(* Logix 5000 project; controller MV vendor 1 type 14 code 217 rev 31.11; software revision 31.00; part 11 of 53 *)
(* tags used below, declared in another part *)
   MC_CIP_String_Result1 : DINT;
   MC_CIP_String_Result2 : DINT;
   MC_CIP_String_Result3 : DINT;
   MC_CIP_String_Result4 : DINT;
   MC_CIP_String_Result5 : DINT;
   MC_CIP_String_Result6 : DINT;
   BH_Draindown_ON : DINT;
   CWD : CHECKWORD_FLAGS;
   FRHR26_31_Valves_ON_Produced : DINT;
   FVHR12_1701 : PlantItem;   // Valve FVHR12_17/01
   FVHR12_1702 : PlantItem;   // Valve FVHR12_17/02
   FVHR12_1703 : PlantItem;   // Valve FVHR12_17/03
   FVHR12_17_Valves_ON : BOOL;   // Check bit to confirm valves for FV12-17 route are open
   FVHR18_21_Valves_ON : BOOL;   // Check bit to confirm valves for FV18-21 route are open
   FVHR18_2501 : PlantItem;   // Valve FVHR18_25/01
   FVHR18_2502 : PlantItem;   // Valve FVHR18_25/02
   FVHR18_2503 : PlantItem;   // Valve FVHR18_25/03
   FVHR18_2504 : PlantItem;   // Valve FVHR18_25/04
   FVHR18_2505 : PlantItem;   // Valve FVHR18_25/05
   FVHR18_2506 : PlantItem;   // Valve FVHR18_25/06
   FVHR1_1101 : PlantItem;   // Valve FVHR1_11/01
   FVHR1_1102 : PlantItem;   // Valve FVHR1_11/02
   FVHR1_1103 : PlantItem;   // Valve FVHR1_11/03
   FVHR1_11_Valves_ON : BOOL;   // Check bit to confirm valves for FV1-11 route are open
   FVHR1_1701 : PlantItem;   // Valve FVHR1_17/01
   FVHR22_25_Valves_ON : BOOL;   // Check bit to confirm valves for FV22-25 route are open
   FVHR26_3101 : PlantItem;   // Valve FVHR26_31/01
   FVHR26_3102 : PlantItem;   // Valve FVHR26_31/02
   FVHR26_3103 : PlantItem;   // Valve FVHR26_31/03
   FVHR26_31_Valves_ON : BOOL;   // Check bit to confirm valves for FV26-31 route are open
   FVHRLTX02_IP : PlantItem;   // Effluent Tank Level Transmitter
   FVHRM02 : PlantItem;   // Valve FVHRM02
   FVHRM03 : PlantItem;   // Valve FVHRM03
   FVHRM04 : PlantItem;   // Valve FVHRM04
   FVHRMD01 : PlantItem;   // Valve FVHRMD01
   FVHRTM01_IP : PlantItem;   // Turbidty Meter FVHRTM01
   IGI_TestBit : BOOL;
   MC_bit_returned : BOOL;
   MC_CH2_CIP_BYPASS_Conditions : BOOL;
   MC_CH2_CIP_BYPASS_DrainConditions : BOOL;
   MC_CH2_CIP_Messages : STRING[20];   // CH2 CIP Scada Messages
   MC_CH2_CIP_YST_Scb_Bypass : BOOL;
   MC_CH2_DR1 : PlantItem;   // CH2_DR1
   MC_CH2_DR2 : PlantItem;   // CH2_DR2
   MC_CH2_DT1 : PlantItem;   // CH2_DT1
   MC_CH2_DT2 : PlantItem;   // CH2_DT2
   MC_CH2_FVBypass_Flush_ALARM : ALARM_DIGITAL;
   MC_CH2_FVBYPASS_H2O_Flush : BOOL;
   MC_CH2_R1 : PlantItem;   // CH2_R1
   MC_CH2_R1R : PlantItem;   // CH2_R1R
   MC_CH2_R2 : PlantItem;   // CH2_R2
   MC_CH2_R2R : PlantItem;   // CH2_R2R
   MC_CH2_R3 : PlantItem;   // CH2_R3
   MC_CH2_R3R : PlantItem;   // CH2_R3R
   MC_CH2_R4 : PlantItem;   // CH2_R4
   MC_CH2_R4R : PlantItem;   // CH2_R4R
   MC_CH2_R5 : PlantItem;   // CH2_R5
   MC_CH2_R5R : PlantItem;   // CH2_R5R
   MC_CH2_R6 : PlantItem;   // CH2_R6
   MC_CH2_R6R : PlantItem;   // CH2_R6R
   MC_CH2_TURBID_High : BOOL;
   MC_CIP_CH2_String_OK : BOOL;
   MC_CIP_CH2_Strings_HopRinse : STRING[30];
   MC_CIP_EFFTank_Full : BOOL;
   MC_CIP_EFFTank_Start_Lvl_Ok : BOOL;
   MC_N10 : INT[255];   // SETTINGS
   MC_N112 : INT[255];   // FVR DATA Data read from FV ro uting PLC
   MC_N113 : INT[255];   // MVR DATA Data read from MV ro uting PLC
   MC_N114 : INT[255];   // YP DATA
   MC_N120 : INT[255];   // C2 PLC Channel 2 PLC data
   MC_N122 : INT[255];   // CH2 PROG Channel 2 CIP progra m
   MC_N200 : INT[255];   // CHK_WORK Plant item fault che cking work area
   MC_N7 : INT[255];   // INTEGER
   MC_P2 : PlantItem;   // P2
   MC_PX_100 : PlantItem;   // PX_100
   MC_PX_101 : PlantItem;   // PX_101
   MC_T125 : TIMER[255];   // CH2 TIMERS Channel 2 timers
   MC_T4 : TIMER[255];   // TIMER
(* MC_Common, continued *)

ROUTINE MC_CH2_GLOBL_125   (* ladder *)
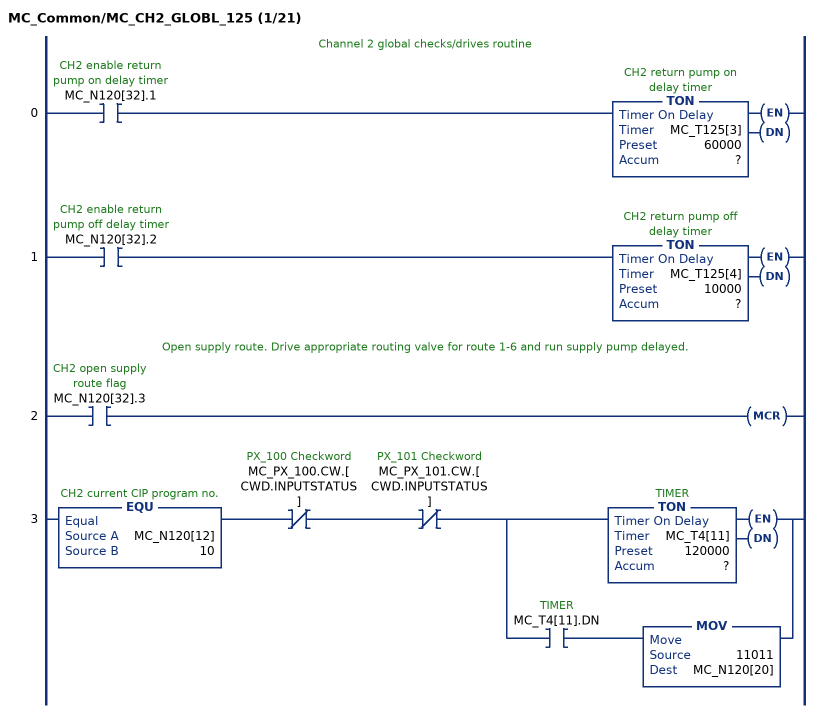
   // Channel 2 global checks/drives routine
   0: XIC(MC_N120[32].1)TON(MC_T125[3],?,?);
   1: XIC(MC_N120[32].2)TON(MC_T125[4],?,?);
   // Open supply route. Drive appropriate routing valve for route 1-6 and run supply pump delayed.
   2: XIC(MC_N120[32].3)MCR();
   3: EQU(MC_N120[12],10)XIO(MC_PX_100.CW.[CWD.INPUTSTATUS])XIO(MC_PX_101.CW.[CWD.INPUTSTATUS])[TON(MC_T4[11],?,?) ,XIC(MC_T4[11].DN) MOV(11011,MC_N120[20]) ];
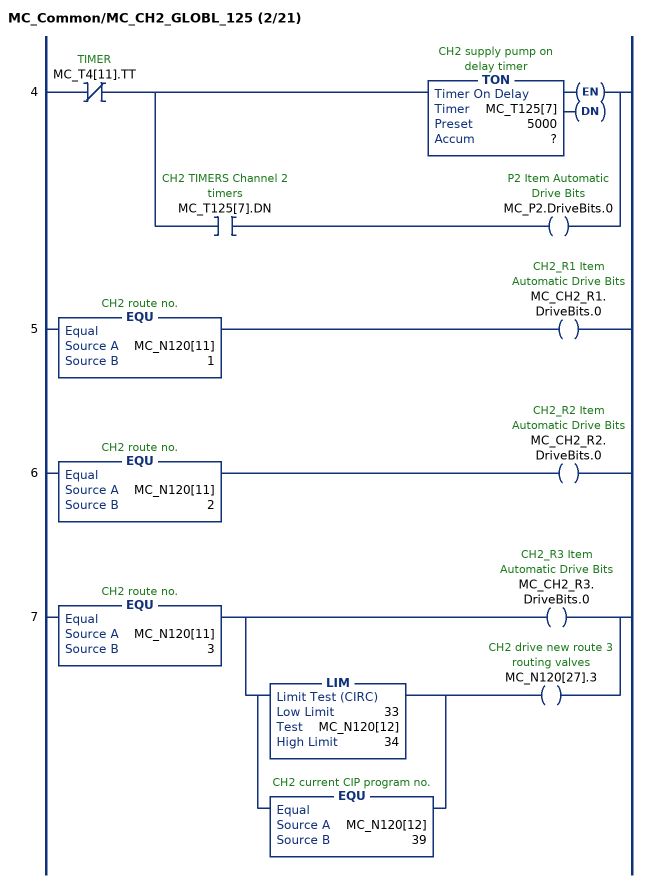
   4: XIO(MC_T4[11].TT)[TON(MC_T125[7],?,?) ,XIC(MC_T125[7].DN) OTE(MC_P2.DriveBits.0) ];
   5: EQU(MC_N120[11],1)OTE(MC_CH2_R1.DriveBits.0);
   6: EQU(MC_N120[11],2)OTE(MC_CH2_R2.DriveBits.0);
   7: EQU(MC_N120[11],3)[OTE(MC_CH2_R3.DriveBits.0) ,[LIM(33,MC_N120[12],34) ,EQU(MC_N120[12],39) ] OTE(MC_N120[27].3) ];
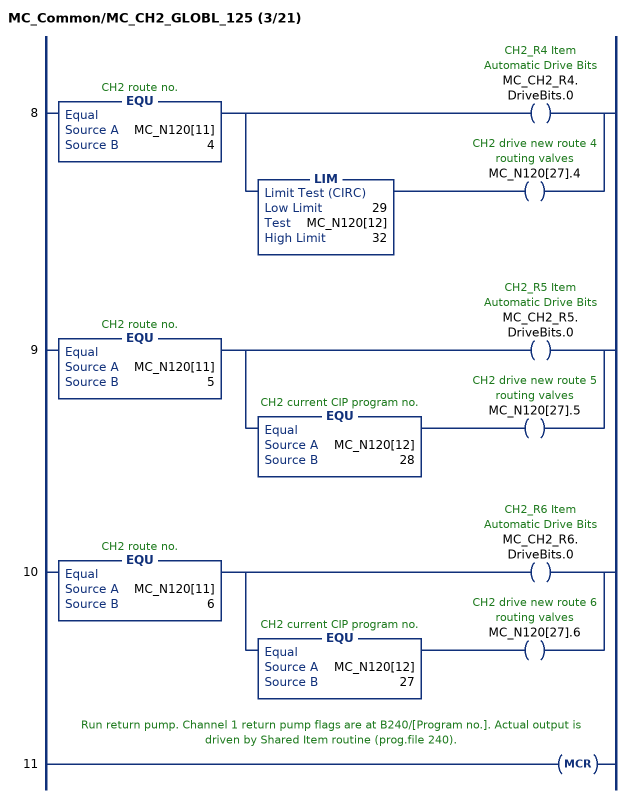
   8: EQU(MC_N120[11],4)[OTE(MC_CH2_R4.DriveBits.0) ,LIM(29,MC_N120[12],32) OTE(MC_N120[27].4) ];
   9: EQU(MC_N120[11],5)[OTE(MC_CH2_R5.DriveBits.0) ,EQU(MC_N120[12],28) OTE(MC_N120[27].5) ];
   10: EQU(MC_N120[11],6)[OTE(MC_CH2_R6.DriveBits.0) ,EQU(MC_N120[12],27) OTE(MC_N120[27].6) ];
   // Run return pump. Channel 1 return pump flags are at B240/[Program no.]. Actual output is driven by Shared Item routine (prog.file 240).
   11: MCR();
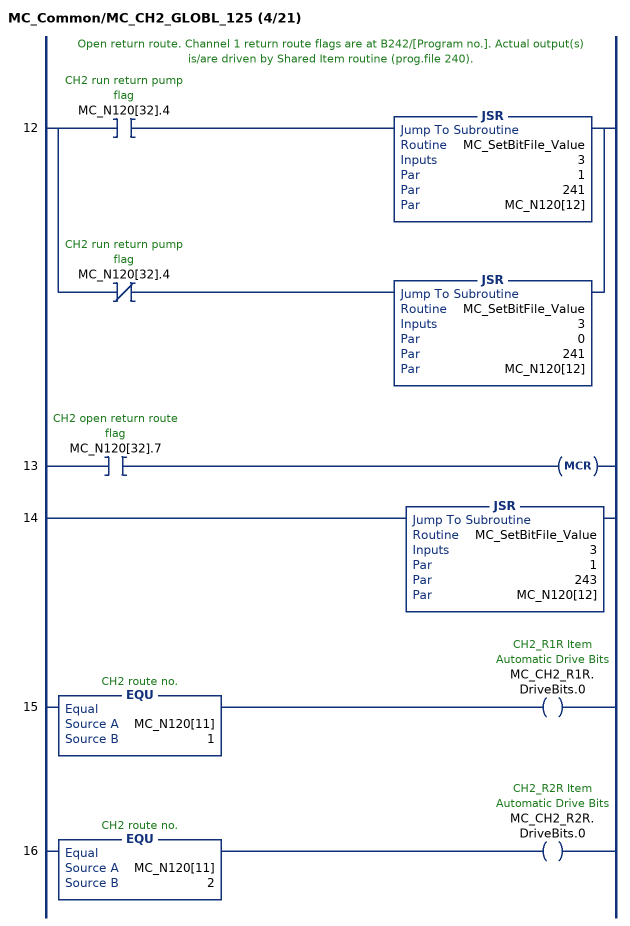
   // Open return route. Channel 1 return route flags are at B242/[Program no.]. Actual output(s) is/are driven by Shared Item routine (prog.file 240).
   12: [XIC(MC_N120[32].4) JSR(MC_SetBitFile_Value,3,1,241,MC_N120[12]) ,XIO(MC_N120[32].4) JSR(MC_SetBitFile_Value,3,0,241,MC_N120[12]) ];
   13: XIC(MC_N120[32].7)MCR();
   14: JSR(MC_SetBitFile_Value,3,1,243,MC_N120[12]);
   15: EQU(MC_N120[11],1)OTE(MC_CH2_R1R.DriveBits.0);
   16: EQU(MC_N120[11],2)OTE(MC_CH2_R2R.DriveBits.0);
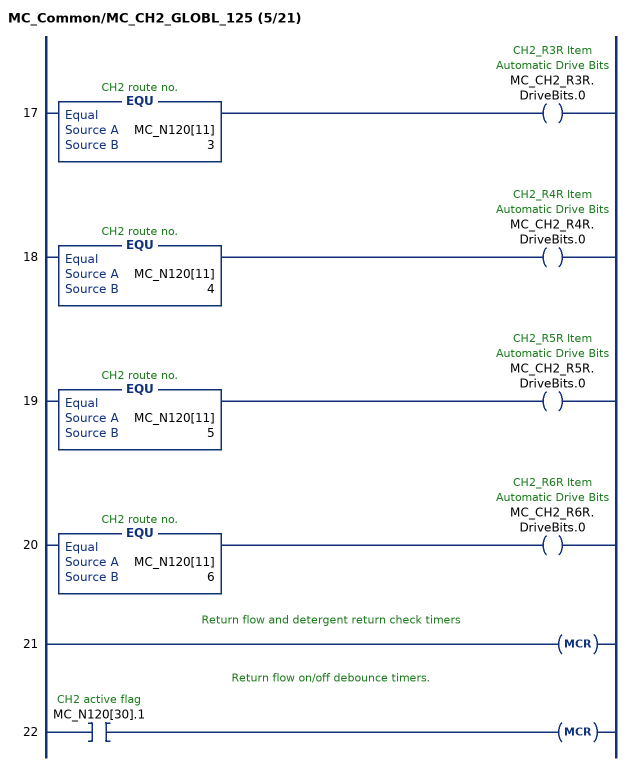
   17: EQU(MC_N120[11],3)OTE(MC_CH2_R3R.DriveBits.0);
   18: EQU(MC_N120[11],4)OTE(MC_CH2_R4R.DriveBits.0);
   19: EQU(MC_N120[11],5)OTE(MC_CH2_R5R.DriveBits.0);
   20: EQU(MC_N120[11],6)OTE(MC_CH2_R6R.DriveBits.0);
   // Return flow and detergent return check timers
   21: MCR();
   // Return flow on/off debounce timers.
   22: XIC(MC_N120[30].1)MCR();
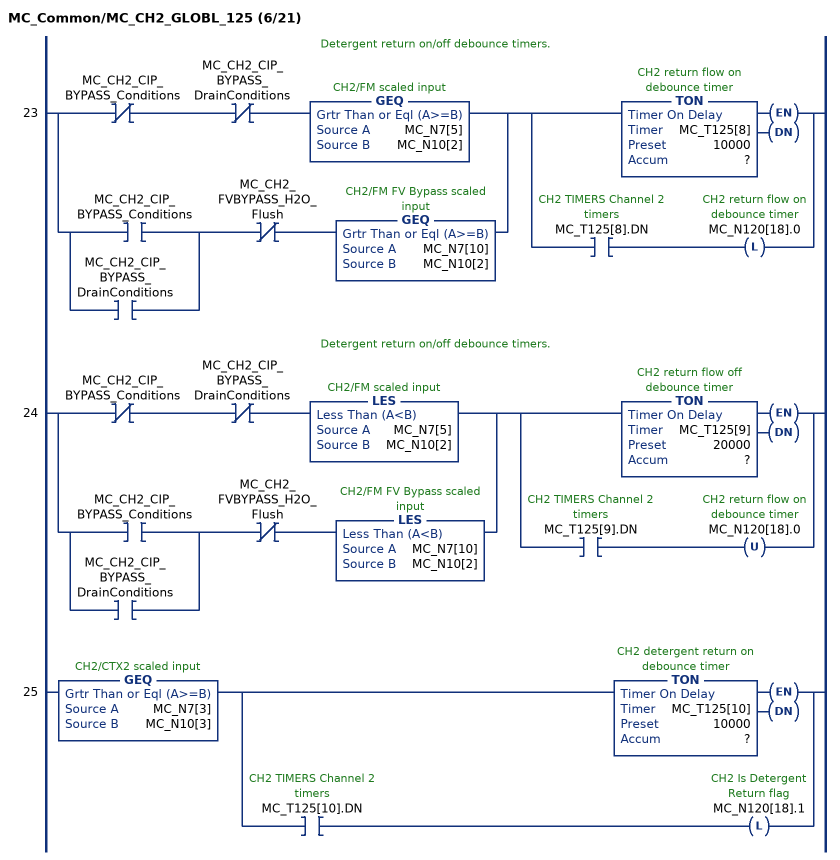
   // Detergent return on/off debounce timers.
   23: [XIO(MC_CH2_CIP_BYPASS_Conditions) XIO(MC_CH2_CIP_BYPASS_DrainConditions) GEQ(MC_N7[5],MC_N10[2]) ,[XIC(MC_CH2_CIP_BYPASS_Conditions) ,XIC(MC_CH2_CIP_BYPASS_DrainConditions) ] XIO(MC_CH2_FVBYPASS_H2O_Flush) GEQ(MC_N7[10],MC_N10[2]) ][TON(MC_T125[8],?,?) ,XIC(MC_T125[8].DN) OTL(MC_N120[18].0) ];
   // Detergent return on/off debounce timers.
   24: [XIO(MC_CH2_CIP_BYPASS_Conditions) XIO(MC_CH2_CIP_BYPASS_DrainConditions) LES(MC_N7[5],MC_N10[2]) ,[XIC(MC_CH2_CIP_BYPASS_Conditions) ,XIC(MC_CH2_CIP_BYPASS_DrainConditions) ] XIO(MC_CH2_FVBYPASS_H2O_Flush) LES(MC_N7[10],MC_N10[2]) ][TON(MC_T125[9],?,?) ,XIC(MC_T125[9].DN) OTU(MC_N120[18].0) ];
   25: GEQ(MC_N7[3],MC_N10[3])[TON(MC_T125[10],?,?) ,XIC(MC_T125[10].DN) OTL(MC_N120[18].1) ];
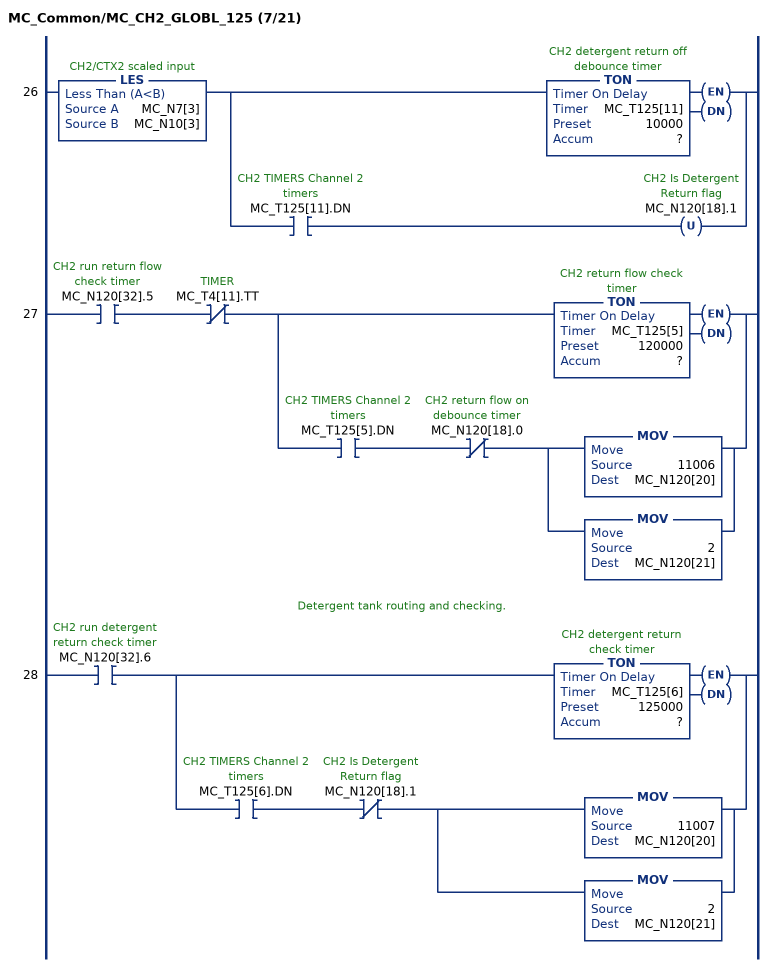
   26: LES(MC_N7[3],MC_N10[3])[TON(MC_T125[11],?,?) ,XIC(MC_T125[11].DN) OTU(MC_N120[18].1) ];
   27: XIC(MC_N120[32].5)XIO(MC_T4[11].TT)[TON(MC_T125[5],?,?) ,XIC(MC_T125[5].DN) XIO(MC_N120[18].0) [MOV(11006,MC_N120[20]) ,MOV(2,MC_N120[21]) ] ];
   // Detergent tank routing and checking.
   28: XIC(MC_N120[32].6)[TON(MC_T125[6],?,?) ,XIC(MC_T125[6].DN) XIO(MC_N120[18].1) [MOV(11007,MC_N120[20]) ,MOV(2,MC_N120[21]) ] ];
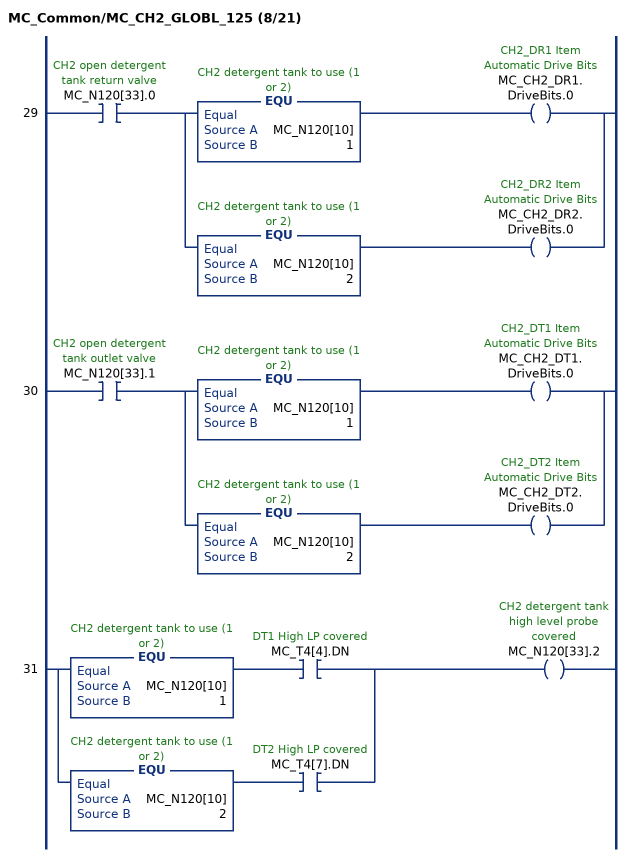
   29: XIC(MC_N120[33].0)[EQU(MC_N120[10],1) OTE(MC_CH2_DR1.DriveBits.0) ,EQU(MC_N120[10],2) OTE(MC_CH2_DR2.DriveBits.0) ];
   30: XIC(MC_N120[33].1)[EQU(MC_N120[10],1) OTE(MC_CH2_DT1.DriveBits.0) ,EQU(MC_N120[10],2) OTE(MC_CH2_DT2.DriveBits.0) ];
   31: [EQU(MC_N120[10],1) XIC(MC_T4[4].DN) ,EQU(MC_N120[10],2) XIC(MC_T4[7].DN) ]OTE(MC_N120[33].2);
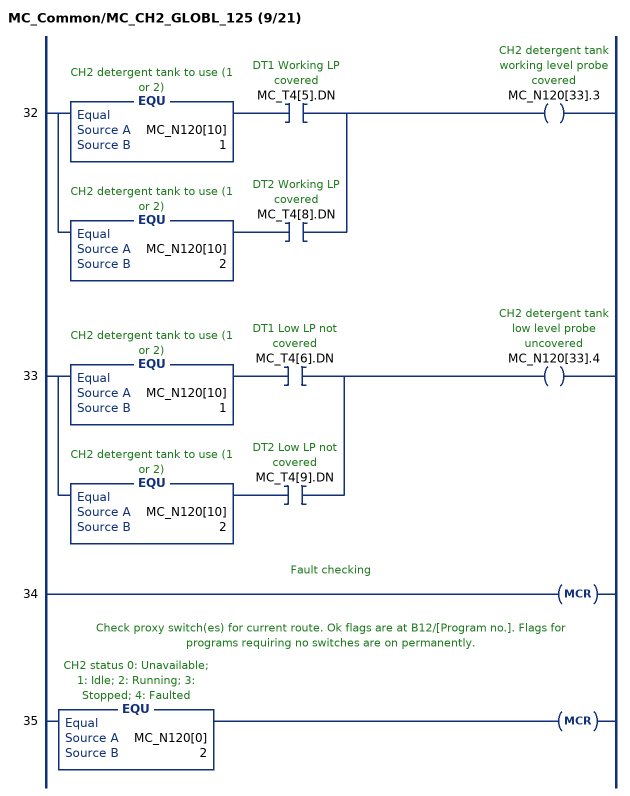
   32: [EQU(MC_N120[10],1) XIC(MC_T4[5].DN) ,EQU(MC_N120[10],2) XIC(MC_T4[8].DN) ]OTE(MC_N120[33].3);
   33: [EQU(MC_N120[10],1) XIC(MC_T4[6].DN) ,EQU(MC_N120[10],2) XIC(MC_T4[9].DN) ]OTE(MC_N120[33].4);
   // Fault checking
   34: MCR();
   // Check proxy switch(es) for current route. Ok flags are at B12/[Program no.]. Flags for programs requiring no switches are on permanently.
   35: EQU(MC_N120[0],2)MCR();
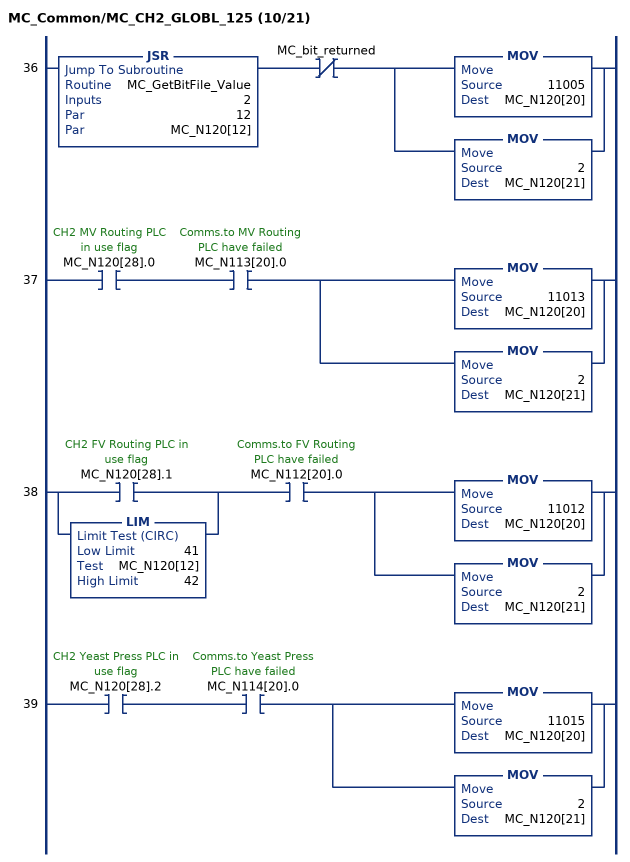
   36: JSR(MC_GetBitFile_Value,2,12,MC_N120[12])XIO(MC_bit_returned)[MOV(11005,MC_N120[20]) ,MOV(2,MC_N120[21]) ];
   37: XIC(MC_N120[28].0)XIC(MC_N113[20].0)[MOV(11013,MC_N120[20]) ,MOV(2,MC_N120[21]) ];
   38: [XIC(MC_N120[28].1) ,LIM(41,MC_N120[12],42) ]XIC(MC_N112[20].0)[MOV(11012,MC_N120[20]) ,MOV(2,MC_N120[21]) ];
   39: XIC(MC_N120[28].2)XIC(MC_N114[20].0)[MOV(11015,MC_N120[20]) ,MOV(2,MC_N120[21]) ];
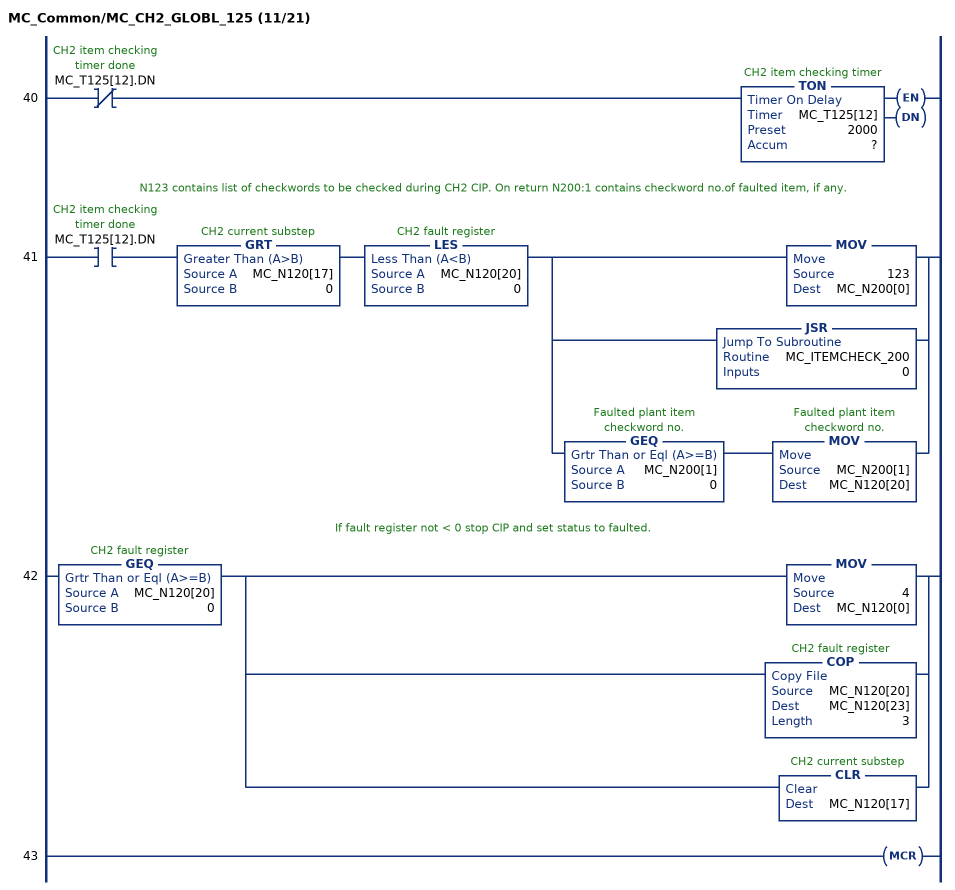
   40: XIO(MC_T125[12].DN)TON(MC_T125[12],?,?);
   // N123 contains list of checkwords to be checked during CH2 CIP. On return N200:1 contains checkword no.of faulted item, if any.
   41: XIC(MC_T125[12].DN)GRT(MC_N120[17],0)LES(MC_N120[20],0)[MOV(123,MC_N200[0]) ,JSR(MC_ITEMCHECK_200,0) ,GEQ(MC_N200[1],0) MOV(MC_N200[1],MC_N120[20]) ];
   // If fault register not < 0 stop CIP and set status to faulted.
   42: GEQ(MC_N120[20],0)[MOV(4,MC_N120[0]) ,COP(MC_N120[20],MC_N120[23],3) ,CLR(MC_N120[17]) ];
   43: MCR();
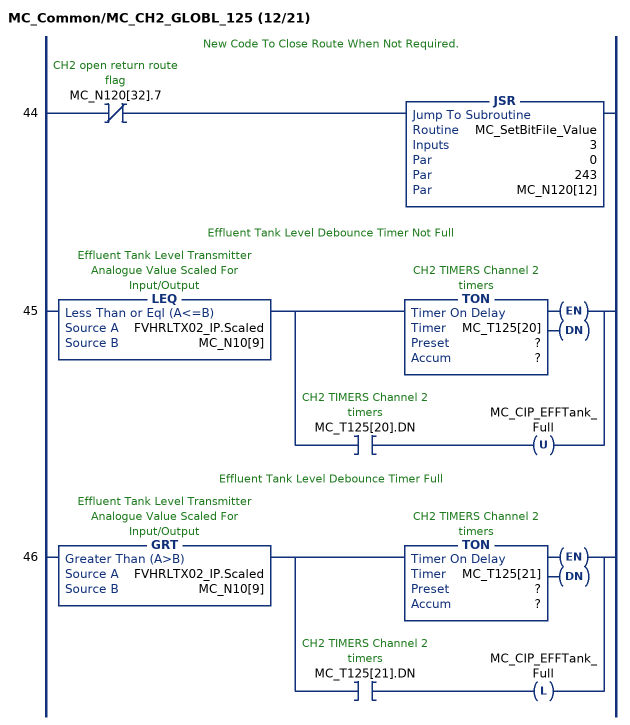
   // New Code To Close Route When Not Required.
   44: XIO(MC_N120[32].7)JSR(MC_SetBitFile_Value,3,0,243,MC_N120[12]);
   // Effluent Tank Level Debounce Timer Not Full
   45: LEQ(FVHRLTX02_IP.Scaled,MC_N10[9])[TON(MC_T125[20],?,?) ,XIC(MC_T125[20].DN) OTU(MC_CIP_EFFTank_Full) ];
   // Effluent Tank Level Debounce Timer Full
   46: GRT(FVHRLTX02_IP.Scaled,MC_N10[9])[TON(MC_T125[21],?,?) ,XIC(MC_T125[21].DN) OTL(MC_CIP_EFFTank_Full) ];
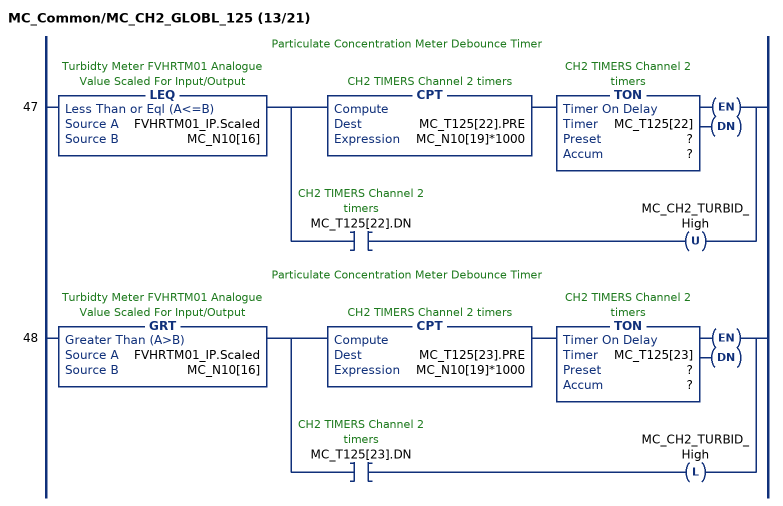
   // Particulate Concentration Meter Debounce Timer
   47: LEQ(FVHRTM01_IP.Scaled,MC_N10[16])[CPT(MC_T125[22].PRE,MC_N10[19]*1000) TON(MC_T125[22],?,?) ,XIC(MC_T125[22].DN) OTU(MC_CH2_TURBID_High) ];
   // Particulate Concentration Meter Debounce Timer
   48: GRT(FVHRTM01_IP.Scaled,MC_N10[16])[CPT(MC_T125[23].PRE,MC_N10[19]*1000) TON(MC_T125[23],?,?) ,XIC(MC_T125[23].DN) OTL(MC_CH2_TURBID_High) ];
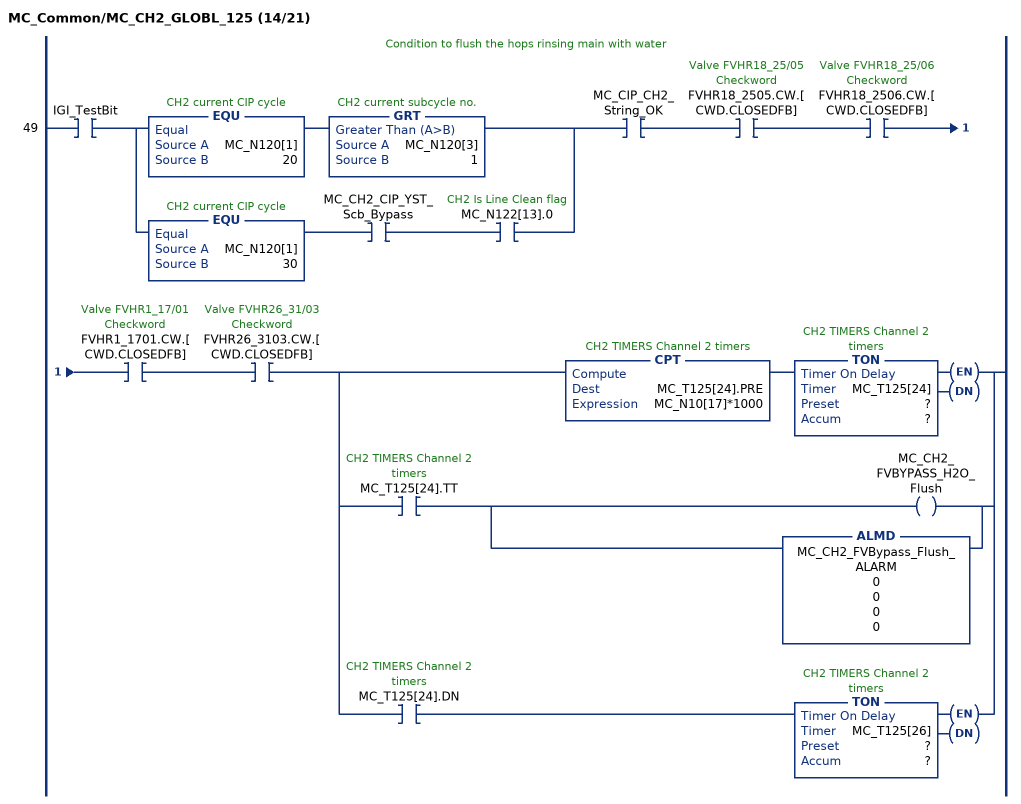
   // Condition to flush the hops rinsing main with water
   49: XIC(IGI_TestBit)[EQU(MC_N120[1],20) GRT(MC_N120[3],1) ,EQU(MC_N120[1],30) XIC(MC_CH2_CIP_YST_Scb_Bypass) XIC(MC_N122[13].0) ]XIC(MC_CIP_CH2_String_OK)XIC(FVHR18_2505.CW.[CWD.CLOSEDFB])XIC(FVHR18_2506.CW.[CWD.CLOSEDFB])XIC(FVHR1_1701.CW.[CWD.CLOSEDFB])XIC(FVHR26_3103.CW.[CWD.CLOSEDFB])[CPT(MC_T125[24].PRE,MC_N10[17]*1000) TON(MC_T125[24],?,?) ,XIC(MC_T125[24].TT) [OTE(MC_CH2_FVBYPASS_H2O_Flush) ,ALMD(MC_CH2_FVBypass_Flush_ALARM,0,0,0,0) ] ,XIC(MC_T125[24].DN) TON(MC_T125[26],?,?) ];
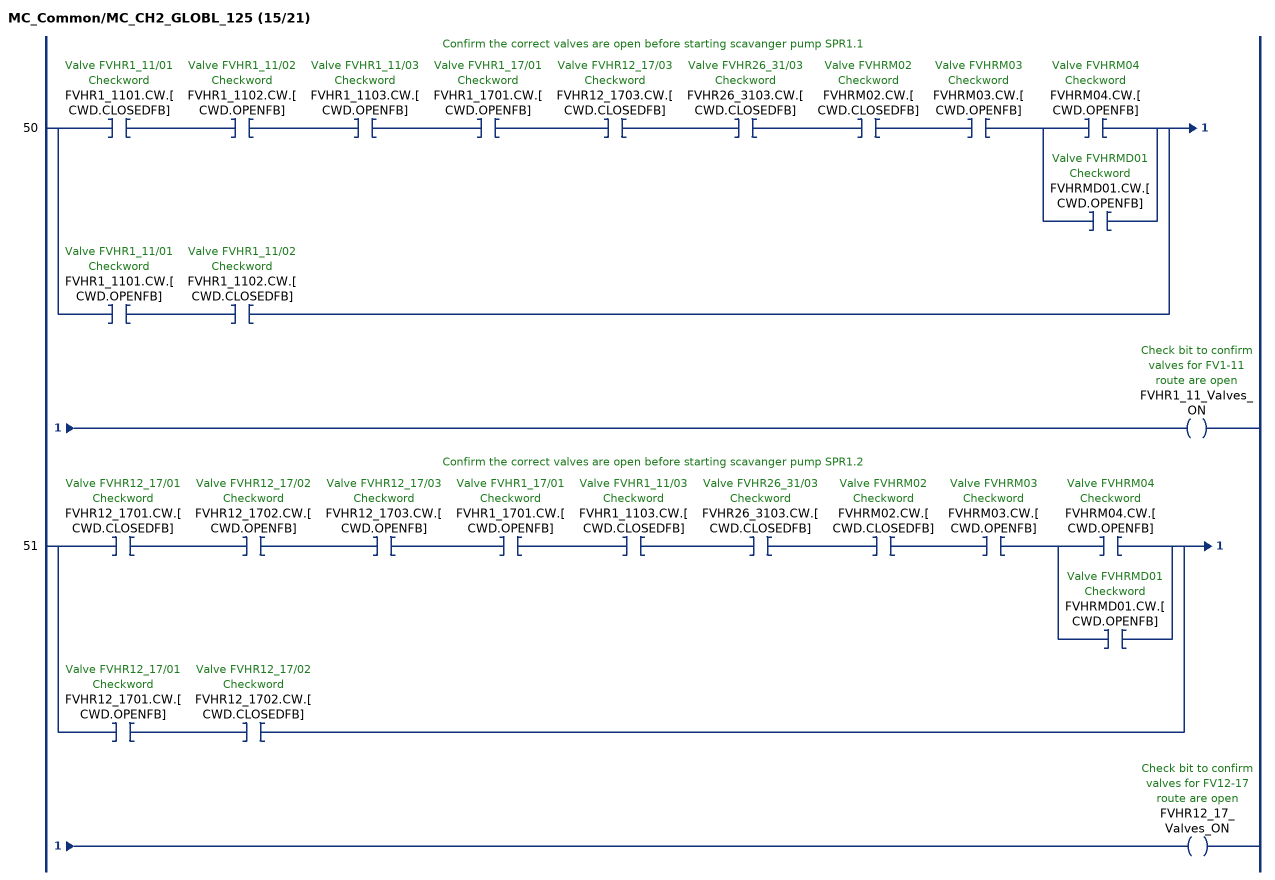
   // Confirm the correct valves are open before starting scavanger pump SPR1.1
   50: [XIC(FVHR1_1101.CW.[CWD.CLOSEDFB]) XIC(FVHR1_1102.CW.[CWD.OPENFB]) XIC(FVHR1_1103.CW.[CWD.OPENFB]) XIC(FVHR1_1701.CW.[CWD.OPENFB]) XIC(FVHR12_1703.CW.[CWD.CLOSEDFB]) XIC(FVHR26_3103.CW.[CWD.CLOSEDFB]) XIC(FVHRM02.CW.[CWD.CLOSEDFB]) XIC(FVHRM03.CW.[CWD.OPENFB]) [XIC(FVHRM04.CW.[CWD.OPENFB]) ,XIC(FVHRMD01.CW.[CWD.OPENFB]) ] ,XIC(FVHR1_1101.CW.[CWD.OPENFB]) XIC(FVHR1_1102.CW.[CWD.CLOSEDFB]) ]OTE(FVHR1_11_Valves_ON);
   // Confirm the correct valves are open before starting scavanger pump SPR1.2
   51: [XIC(FVHR12_1701.CW.[CWD.CLOSEDFB]) XIC(FVHR12_1702.CW.[CWD.OPENFB]) XIC(FVHR12_1703.CW.[CWD.OPENFB]) XIC(FVHR1_1701.CW.[CWD.OPENFB]) XIC(FVHR1_1103.CW.[CWD.CLOSEDFB]) XIC(FVHR26_3103.CW.[CWD.CLOSEDFB]) XIC(FVHRM02.CW.[CWD.CLOSEDFB]) XIC(FVHRM03.CW.[CWD.OPENFB]) [XIC(FVHRM04.CW.[CWD.OPENFB]) ,XIC(FVHRMD01.CW.[CWD.OPENFB]) ] ,XIC(FVHR12_1701.CW.[CWD.OPENFB]) XIC(FVHR12_1702.CW.[CWD.CLOSEDFB]) ]OTE(FVHR12_17_Valves_ON);
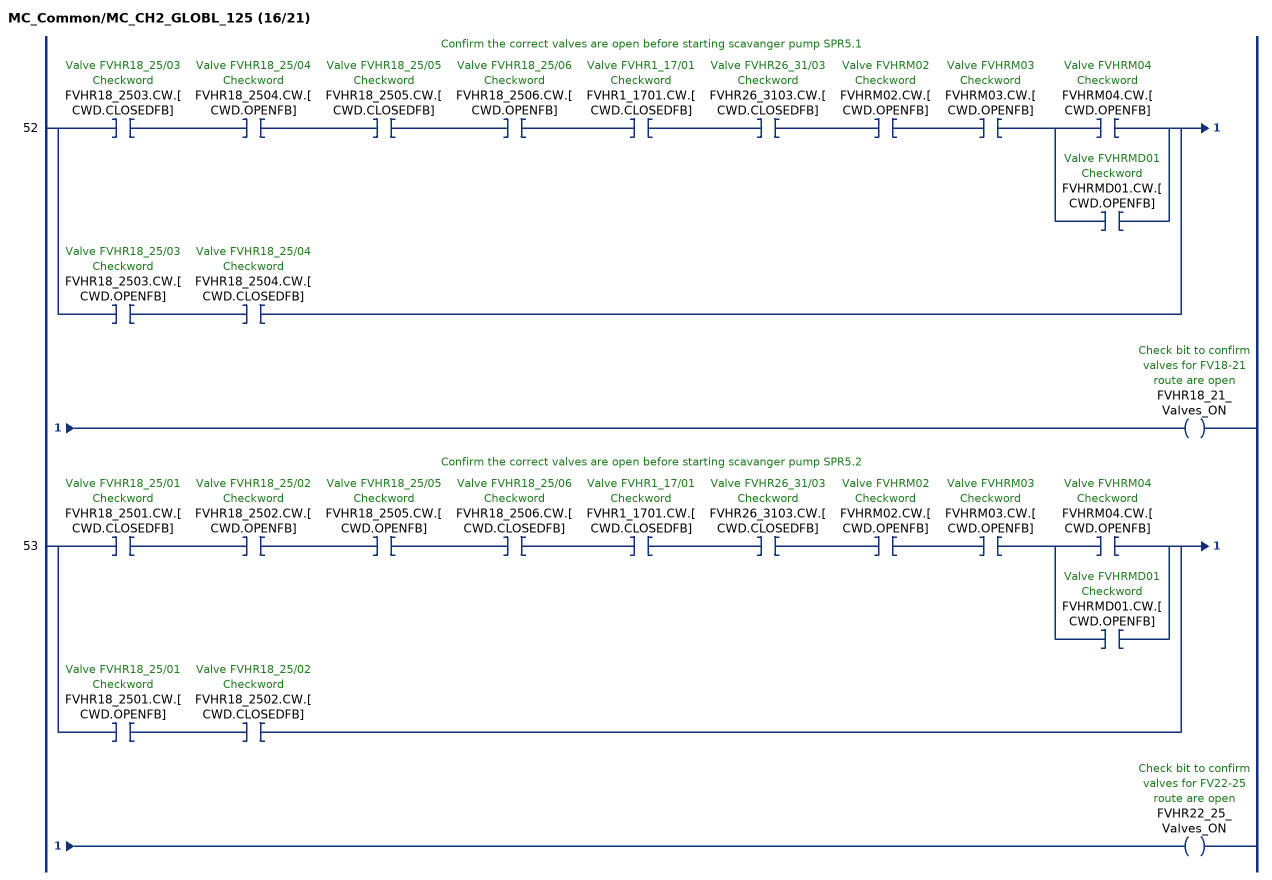
   // Confirm the correct valves are open before starting scavanger pump SPR5.1
   52: [XIC(FVHR18_2503.CW.[CWD.CLOSEDFB]) XIC(FVHR18_2504.CW.[CWD.OPENFB]) XIC(FVHR18_2505.CW.[CWD.CLOSEDFB]) XIC(FVHR18_2506.CW.[CWD.OPENFB]) XIC(FVHR1_1701.CW.[CWD.CLOSEDFB]) XIC(FVHR26_3103.CW.[CWD.CLOSEDFB]) XIC(FVHRM02.CW.[CWD.OPENFB]) XIC(FVHRM03.CW.[CWD.OPENFB]) [XIC(FVHRM04.CW.[CWD.OPENFB]) ,XIC(FVHRMD01.CW.[CWD.OPENFB]) ] ,XIC(FVHR18_2503.CW.[CWD.OPENFB]) XIC(FVHR18_2504.CW.[CWD.CLOSEDFB]) ]OTE(FVHR18_21_Valves_ON);
   // Confirm the correct valves are open before starting scavanger pump SPR5.2
   53: [XIC(FVHR18_2501.CW.[CWD.CLOSEDFB]) XIC(FVHR18_2502.CW.[CWD.OPENFB]) XIC(FVHR18_2505.CW.[CWD.OPENFB]) XIC(FVHR18_2506.CW.[CWD.CLOSEDFB]) XIC(FVHR1_1701.CW.[CWD.CLOSEDFB]) XIC(FVHR26_3103.CW.[CWD.CLOSEDFB]) XIC(FVHRM02.CW.[CWD.OPENFB]) XIC(FVHRM03.CW.[CWD.OPENFB]) [XIC(FVHRM04.CW.[CWD.OPENFB]) ,XIC(FVHRMD01.CW.[CWD.OPENFB]) ] ,XIC(FVHR18_2501.CW.[CWD.OPENFB]) XIC(FVHR18_2502.CW.[CWD.CLOSEDFB]) ]OTE(FVHR22_25_Valves_ON);
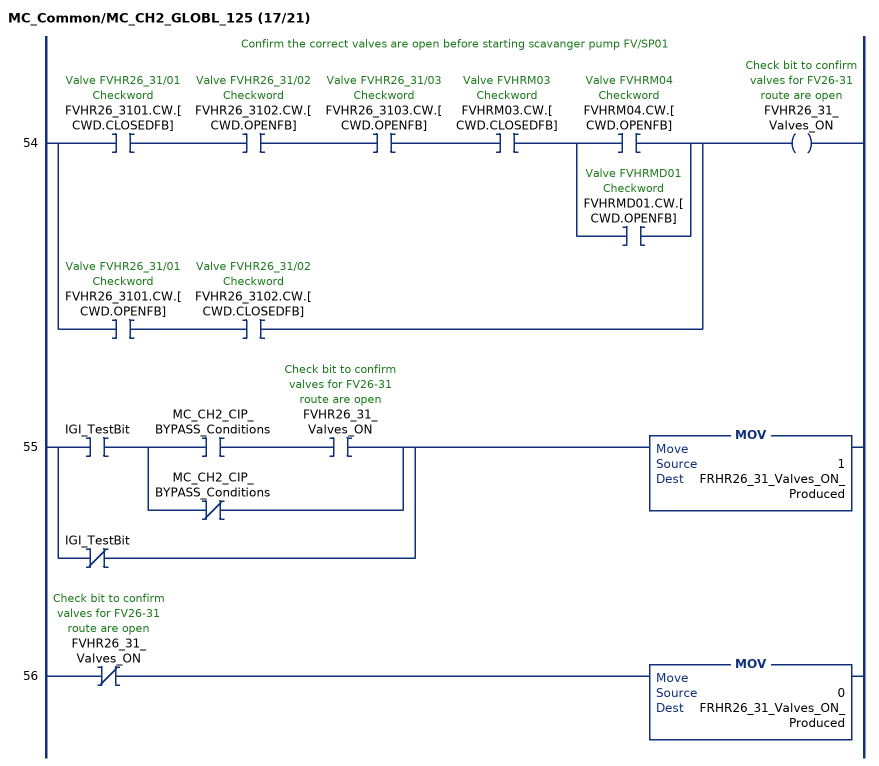
   // Confirm the correct valves are open before starting scavanger pump FV/SP01
   54: [XIC(FVHR26_3101.CW.[CWD.CLOSEDFB]) XIC(FVHR26_3102.CW.[CWD.OPENFB]) XIC(FVHR26_3103.CW.[CWD.OPENFB]) XIC(FVHRM03.CW.[CWD.CLOSEDFB]) [XIC(FVHRM04.CW.[CWD.OPENFB]) ,XIC(FVHRMD01.CW.[CWD.OPENFB]) ] ,XIC(FVHR26_3101.CW.[CWD.OPENFB]) XIC(FVHR26_3102.CW.[CWD.CLOSEDFB]) ]OTE(FVHR26_31_Valves_ON);
   55: [XIC(IGI_TestBit) [XIC(MC_CH2_CIP_BYPASS_Conditions) XIC(FVHR26_31_Valves_ON) ,XIO(MC_CH2_CIP_BYPASS_Conditions) ] ,XIO(IGI_TestBit) ]MOV(1,FRHR26_31_Valves_ON_Produced);
   56: XIO(FVHR26_31_Valves_ON)MOV(0,FRHR26_31_Valves_ON_Produced);
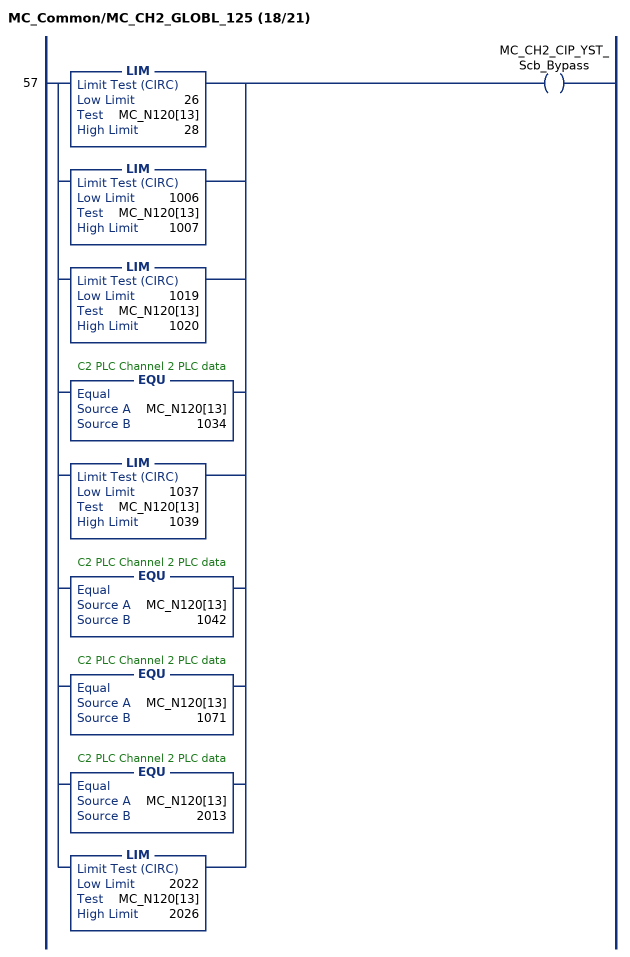
   57: [LIM(26,MC_N120[13],28) ,LIM(1006,MC_N120[13],1007) ,LIM(1019,MC_N120[13],1020) ,EQU(MC_N120[13],1034) ,LIM(1037,MC_N120[13],1039) ,EQU(MC_N120[13],1042) ,EQU(MC_N120[13],1071) ,EQU(MC_N120[13],2013) ,LIM(2022,MC_N120[13],2026) ]OTE(MC_CH2_CIP_YST_Scb_Bypass);
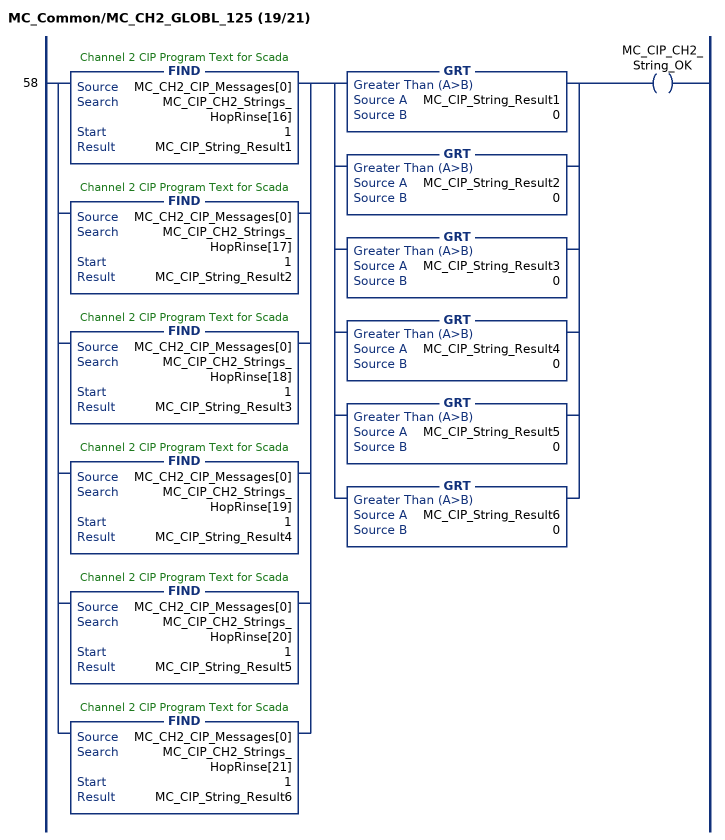
   58: [FIND(MC_CH2_CIP_Messages[0],MC_CIP_CH2_Strings_HopRinse[16],1,MC_CIP_String_Result1) ,FIND(MC_CH2_CIP_Messages[0],MC_CIP_CH2_Strings_HopRinse[17],1,MC_CIP_String_Result2) ,FIND(MC_CH2_CIP_Messages[0],MC_CIP_CH2_Strings_HopRinse[18],1,MC_CIP_String_Result3) ,FIND(MC_CH2_CIP_Messages[0],MC_CIP_CH2_Strings_HopRinse[19],1,MC_CIP_String_Result4) ,FIND(MC_CH2_CIP_Messages[0],MC_CIP_CH2_Strings_HopRinse[20],1,MC_CIP_String_Result5) ,FIND(MC_CH2_CIP_Messages[0],MC_CIP_CH2_Strings_HopRinse[21],1,MC_CIP_String_Result6) ][GRT(MC_CIP_String_Result1,0) ,GRT(MC_CIP_String_Result2,0) ,GRT(MC_CIP_String_Result3,0) ,GRT(MC_CIP_String_Result4,0) ,GRT(MC_CIP_String_Result5,0) ,GRT(MC_CIP_String_Result6,0) ]OTE(MC_CIP_CH2_String_OK);
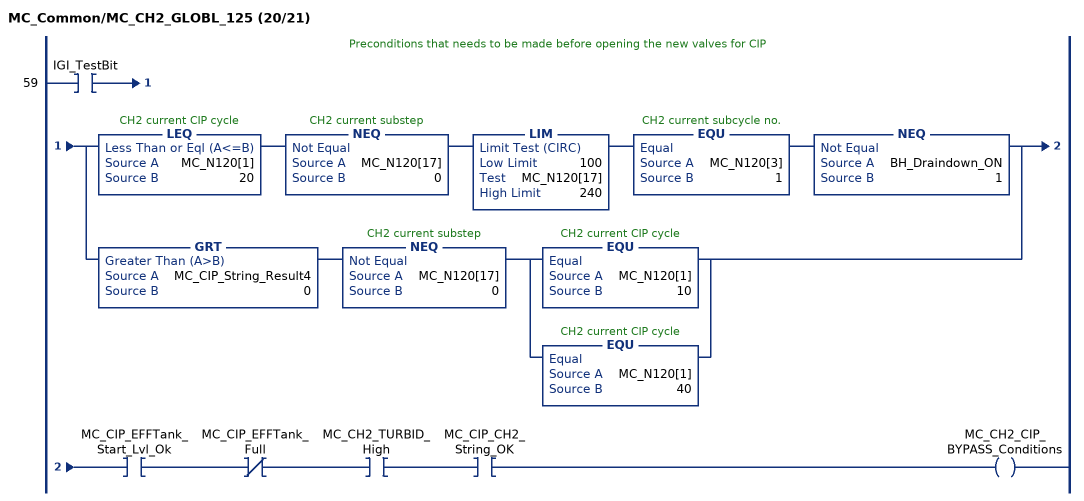
   // Preconditions that needs to be made before opening the new valves for CIP
   59: XIC(IGI_TestBit)[LEQ(MC_N120[1],20) NEQ(MC_N120[17],0) LIM(100,MC_N120[17],240) EQU(MC_N120[3],1) NEQ(BH_Draindown_ON,1) ,GRT(MC_CIP_String_Result4,0) NEQ(MC_N120[17],0) [EQU(MC_N120[1],10) ,EQU(MC_N120[1],40) ] ]XIC(MC_CIP_EFFTank_Start_Lvl_Ok)XIO(MC_CIP_EFFTank_Full)XIC(MC_CH2_TURBID_High)XIC(MC_CIP_CH2_String_OK)OTE(MC_CH2_CIP_BYPASS_Conditions);
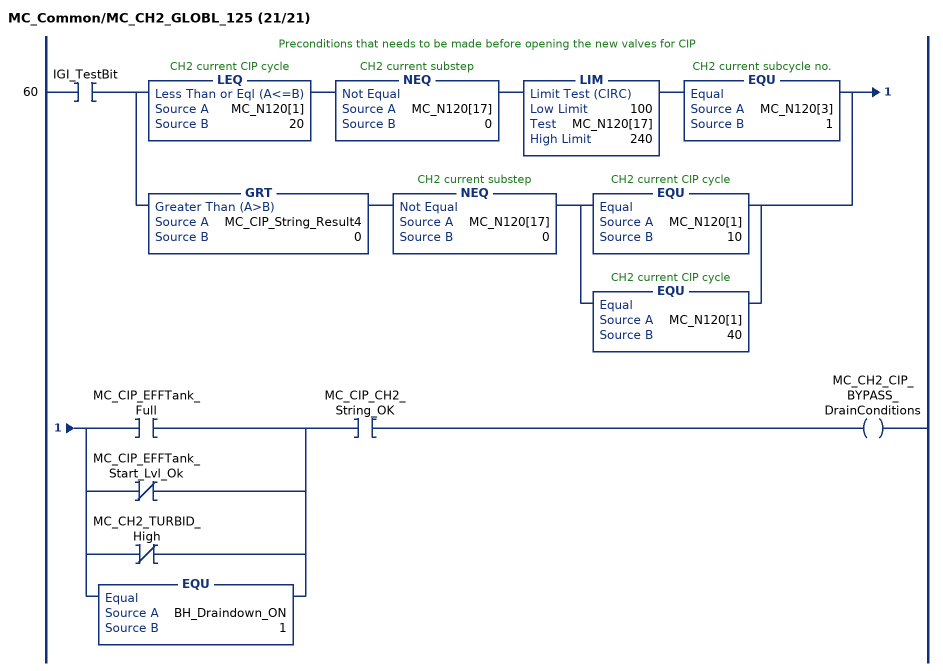
   // Preconditions that needs to be made before opening the new valves for CIP
   60: XIC(IGI_TestBit)[LEQ(MC_N120[1],20) NEQ(MC_N120[17],0) LIM(100,MC_N120[17],240) EQU(MC_N120[3],1) ,GRT(MC_CIP_String_Result4,0) NEQ(MC_N120[17],0) [EQU(MC_N120[1],10) ,EQU(MC_N120[1],40) ] ][XIC(MC_CIP_EFFTank_Full) ,XIO(MC_CIP_EFFTank_Start_Lvl_Ok) ,XIO(MC_CH2_TURBID_High) ,EQU(BH_Draindown_ON,1) ]XIC(MC_CIP_CH2_String_OK)OTE(MC_CH2_CIP_BYPASS_DrainConditions);
END_ROUTINE
